// TIA Portal project "TestEssProtoFreia" (V13)

(* hardware
DEVICE "Station S7300/ET200M_1"  S7-300 station
   slot 0: "Châssis_0"  Rail  6ES7 390-1***0-0AA0
   slot 1: "Châssis_1"  Rail  6ES7 390-1***0-0AA0
   slot 1: "PS 307 2A_1"  PS 307 2A  6ES7 307-1BA01-0AA0
   slot 1: "PS 307 2A_1"  PS 307 2A  6ES7 307-1BA01-0AA0
   slot 2: "PLC_1"  CPU 315-2 DP  6ES7 315-2AH14-0AB0  V3.3
      slot 0: "Interface MPI_1"  MPI
      slot 1: "Interface DP_1"  DP
   slot 3: "IM 360_1"  6ES7 360-3AA01-0AA0
      slot 1: "Interface d'émission IM_1"  6ES7 360-3AA00-0AA0
   slot 3: "IM 361_1"  6ES7 361-3CA01-0AA0
      slot 1: "Interface d'émission IM_1"  6ES7 360-3AA00-0AA0
      slot 2: "Interface de réception IM_1"  6ES7 361-3CA00-0AA0
   slot 4: "DO 16x24VDC/0.5A_2"  DO16 x 24VDC / 0.5A  6ES7 322-1BH01-0AA0
   slot 4: "CP 343-1 Lean_1"  CP 343-1 LEAN  6GK7 343-1CX10-0XE0  V2.2
   slot 5: "DO 16x24VDC/0.5A_1"  DO16 x 24VDC / 0.5A  6ES7 322-1BH01-0AA0
   slot 5: "DI 16x24VDC_1"  DI16 x 24VDC  6ES7 321-1BH02-0AA0
   slot 6: "AI 8x12BIT_1"  AI8 x 12 bits  6ES7 331-7KF02-0AB0
   slot 6: "AI 8x12BIT_1"  AI8 x 12 bits  6ES7 331-7KF02-0AB0
   slot 7: "AI 8x12BIT_2"  AI8 x 12 bits  6ES7 331-7KF02-0AB0
   slot 7: "AO 8x12BIT_1"  AO8 x 12 bits  6ES7 332-5HF00-0AB0
   slot 8: "AI 8x12BIT_3"  AI8 x 12 bits  6ES7 331-7KF02-0AB0
   slot 8: "AO 4x12BIT_1"  AO4 x 12 bits  6ES7 332-5HD01-0AB0
   slot 9: "AI 8x16BIT_1"  AI8 x 16 bits  6ES7 331-7NF00-0AB0
   slot 9: "AO 4x12BIT_2"  AO4 x 12 bits  6ES7 332-5HD01-0AB0
DEVICE "Appareil GSD_1"  GSD.Device
   slot 0: "Châssis_0"  Rail
DEVICE "Appareil GSD_3"  GSD.Device
   slot 0: "Châssis_0"  Rail
DEVICE "Appareil GSD_4"  GSD.Device
   slot 0: "Châssis_0"  Rail
*)

// ===== PLC "PLC_1"  CPU 315-2 DP =====

VAR_GLOBAL   // PLC tag table "Table de variables standard"
   "TT_04" AT %ID720 : Real;
   "TT_218" AT %ID724 : Real;
   "TT_08CM" AT %ID728 : Real;
   "TT_217" AT %ID732 : Real;
   "TT_210" AT %ID736 : Real;
   "TT_209" AT %ID740 : Real;
   "TT_214" AT %ID744 : Real;
   "TT_03" AT %ID780 : Real;
   "TT_205" AT %ID784 : Real;
   "TT_05" AT %ID788 : Real;
   "TT_213" AT %ID792 : Real;
   "TT_14" AT %ID796 : Real;
   "TT_203" AT %ID800 : Real;
   "TT_204" AT %ID804 : Real;
   "TT_211" AT %ID808 : Real;
   "TT_202" AT %ID336 : Real;
   "TT_201" AT %ID340 : Real;
   "TT_104" AT %ID344 : Real;
   "TT_01CM" AT %ID348 : Real;
   "TT_115" AT %ID352 : Real;
   "TT_115bis" AT %ID356 : Real;
   "TT_208" AT %ID360 : Real;
   "TT_07" AT %ID364 : Real;
   "TT_12" AT %ID404 : Real;
   "TT_101" AT %ID408 : Real;
   "TT_103" AT %ID412 : Real;
   "TT_102" AT %ID416 : Real;
   "TT_04bis" AT %ID420 : Real;
   "TT_206" AT %ID424 : Real;
   "TT_02" AT %ID844 : Real;
   "TT_117" AT %ID856 : Real;
   "TT_106" AT %ID860 : Real;
   "TT_116" AT %ID864 : Real;
   "TT_118" AT %ID868 : Real;
   "TT_110" AT %ID872 : Real;
   "TT_207" AT %ID908 : Real;
   "TT_111" AT %ID924 : Real;
   "TT_107" AT %ID928 : Real;
   "TT_06" AT %ID932 : Real;
   "Tag_1" AT %IW3 : Word;
   "TimerDefauCom1" AT %T20 : Timer;
   "TimerDefauCom2" AT %T21 : Timer;
   "TT_215" AT %ID716 : Real;
   "CABTF4_voie10" AT %ID912 : Real;
   "CABTF4_voie11" AT %ID916 : Real;
   "CABTF4_voie12" AT %ID920 : Real;
   "Tag_45" AT %MD224 : Real;
   "Tag_46" AT %MW230 : Word;
   "Tag_47" AT %MW240 : Word;
   "Tag_48" AT %MD240 : Real;
   "Tag_49" AT %MD238 : DWord;
   "Tag_50" AT %MW238 : Word;
   "Tag_51" AT %MW242 : Word;
   "Tag_52" AT %MD244 : Real;
   "Tag_53" AT %IW388 : Int;
   "Tag_27" AT %MW600 : Word;
   "Tag_28" AT %MD602 : Real;
   "Tag_30" AT %M700.0 : Bool;
   "Tag_31" AT %M700.1 : Bool;
   "Tag_32" AT %M800.0 : Bool;
   "Tag_34" AT %MW804 : Int;
   "Tag_36" AT %MD808 : Real;
   "Tag_37" AT %MD812 : Real;
   "Tag_38" AT %MW816 : Word;
   "Tag_40" AT %M800.1 : Bool;
   "Tag_41" AT %M800.2 : Bool;
   "Tag_42" AT %MW802 : Int;
   "Tag_43" AT %MD804 : Real;
   "Tag_54" AT %MW820 : Word;
   "TT103_OHM" AT %MD820 : Real;
   "Tag_56" AT %IW646 : Word;
   "Tag_57" AT %IW648 : Word;
   "Tag_58" AT %IW480 : Word;
   "Tag_59" AT %IW482 : Word;
   "Tag_60" AT %IW472 : Word;
   "Tag_61" AT %IW474 : Word;
   "Tag_62" AT %IW464 : Word;
   "Tag_63" AT %IW466 : Word;
   "LocalMode" AT %M251.0 : Bool;
   "Tag_3" AT %M3.6 : Bool;
END_VAR

VAR_GLOBAL   // PLC tag table "Digital Input"
   "GV_70_CmInsulVacc:Open" AT %I0.0 : Bool;   // Cryomodule insulating vacuum Gate valve 70 open
   "GV_70_CmInsulVacc:Close" AT %I0.1 : Bool;   // Cryomodule insulating vacuum Gate valve 70 close
   "GV_71_CmInsulVacc:Open" AT %I0.3 : Bool;   // Cryomodule insulating vacuum Gate valve 71 open
   "GV_71_CmInsulVacc:Close" AT %I0.4 : Bool;   // Cryomodule insulating vacuum Gate valve 71 close
   "GV_72_VbInsulVacc:Open" AT %I0.6 : Bool;   // Cryomodule insulating vacuum Gate valve 72 open
   "GV_72_VbInsulVacc:Close" AT %I0.7 : Bool;   // Cryomodule insulating vacuum Gate valve 72 close
   "GV72_closed" AT %I1.1 : Bool;   // Cryomodule insulating vacuum Gate valve 72 closed
   "GV70_open" AT %I1.2 : Bool;   // Cryomodule insulating vacuum Gate valve 70 open
   "Tag_4" AT %I2.0 : Bool;
   "GV72_open" AT %I1.0 : Bool;   // Cryomodule insulating vacuum Gate valve 72 open
   "GV70_closed" AT %I1.3 : Bool;   // Cryomodule insulating vacuum Gate valve 70 closed
   "RV90_open" AT %I1.4 : Bool;   // He release valve
   "RV90_closed" AT %I1.5 : Bool;   // He release valve
END_VAR

VAR_GLOBAL   // PLC tag table "analog output"
   "CMD_CV_01" AT %QW384 : Int;
   "CMD_CV_02" AT %QW386 : Int;
   "CMD_CV_03" AT %QW388 : Int;
   "CMD_CV_04" AT %QW390 : Int;
   "CMD_CV_05" AT %QW392 : Int;
   "CMD_CV_07" AT %QW394 : Int;
   "CMD_CV_60" AT %QW396 : Int;
   "CMD_CV_61" AT %QW398 : Int;
   "CMD_CV_62" AT %QW400 : Int;
   "Sana_ASCO_1" AT %QW402 : Int;
   "Sana_ASCO_2" AT %QW404 : Int;
END_VAR

VAR_GLOBAL   // PLC tag table "mem"
   "always_1" AT %M0.1 : Bool;
   "always_0" AT %M0.0 : Bool;
   "unscal_ret_val" AT %MW40 : Word;
   "CV01_HMI_VAL" AT %MD4 : Real;
   "CV02_HMI_VAL" AT %MD8 : Real;
   "CV03_HMI_VAL" AT %MD12 : Real;
   "CV04_HMI_VAL" AT %MD16 : Real;
   "CV05_HMI_VAL" AT %MD20 : Real;
   "CV07_HMI_VAL" AT %MD24 : Real;
   "CV60_HMI_VAL" AT %MD28 : Real;
   "CV61_HMI_VAL" AT %MD36 : Real;
   "unscal_ret_val_1" AT %MW42 : Word;
   "unscal_ret_val_2" AT %MW44 : Word;
   "unscal_ret_val_3" AT %MW46 : Word;
   "unscal_ret_val_4" AT %MW48 : Word;
   "unscal_ret_val_5" AT %MW50 : Word;
   "unscal_ret_val_6" AT %MW52 : Word;
   "unscal_ret_val_7" AT %MW54 : Word;
   "unscal_ret_val_8" AT %MW56 : Word;
   "CV62_HMI_VAL" AT %MD32 : Real;
   "Tag_7" AT %MD701 : Real;
   "Tag_8" AT %MD706 : Real;
   "Tag_9" AT %MD710 : Real;
   "Tag_10" AT %MD714 : Real;
   "Tag_11" AT %MD718 : Real;
   "Tag_12" AT %MD722 : Real;
   "Tag_13" AT %MD726 : Real;
   "Tag_14" AT %MD730 : Real;
   "Tag_15" AT %MD734 : Real;
   "Tag_16" AT %MW100 : Word;
   "Tag_17" AT %MW102 : Word;
   "Tag_18" AT %MW104 : Word;
   "Tag_19" AT %MW106 : Word;
   "Tag_20" AT %MW108 : Word;
   "Tag_21" AT %MW110 : Word;
   "Tag_22" AT %MW112 : Word;
   "Tag_23" AT %MW114 : Word;
   "Tag_24" AT %MW116 : Word;
   "TT670_(OHMS)" AT %MD58 : Real;
   "LT03_DepHaut" AT %M0.3 : Bool;
   "LT03_DepBas" AT %M0.4 : Bool;
   "LT03_DefSond" AT %M0.5 : Bool;
   "LT03_TypeDef" AT %MW66 : Int;
   "LT03_ValMax" AT %MD72 : Real;
   "LT03_ValMin" AT %MD76 : Real;
   "LT03_NiveauHel" AT %MD80 : Real;
   "CV02_ManAuto" AT %M0.6 : Bool;
   "CV03_ManAuto" AT %M0.7 : Bool;
   "CV61_ManAuto" AT %M1.0 : Bool;
   "ScaleErreurPT60" AT %MW68 : Word;
   "ScaleErreurPT01" AT %MW88 : Word;
   "ScaleErreurVidePT73" AT %MW90 : Word;
   "VidePT73Tension" AT %MD92 : Real;
   "CV01PosInit" AT %M1.1 : Bool;
   "CV02PosInit" AT %M1.2 : Bool;
   "CV03PosInit" AT %M1.3 : Bool;
   "CV04PosInit" AT %M1.4 : Bool;
   "CV05PosInit" AT %M1.5 : Bool;
   "CV07PosInit" AT %M1.6 : Bool;
   "CV60PosInit" AT %M1.7 : Bool;
   "CV61PosInit" AT %M62.0 : Bool;
   "CV62PosInit" AT %M62.1 : Bool;
   "CmdVanneEtatInitial" AT %M62.2 : Bool;
   "VanneEnPositionInitial" AT %M62.3 : Bool;
   "CmdVanneEtatCdt" AT %M62.4 : Bool;
   "Etat initial" AT %M62.5 : Bool;
   "CV01PosCdt" AT %M62.6 : Bool;
   "CV02PosCdt" AT %M62.7 : Bool;
   "CV03PosCdt" AT %M63.0 : Bool;
   "CV04PosCdt" AT %M63.1 : Bool;
   "CV05PosCdt" AT %M63.2 : Bool;
   "CV07PosCdt" AT %M63.3 : Bool;
   "CV60PosCdt" AT %M63.4 : Bool;
   "CV61PosCdt" AT %M63.5 : Bool;
   "CV62PosCdt" AT %M63.6 : Bool;
   "VanneEnPositionCdt" AT %M63.7 : Bool;
   "EtatCdtCryo" AT %M64.0 : Bool;
   "ScaleErreurVidePT71" AT %MW96 : Word;
   "VidePT71Tension" AT %MD118 : Real;
   "AutorizationMefAzote" AT %M64.1 : Bool;
   "ReguleCV61ON" AT %M64.2 : Bool;
   "CmdVanneEtatMEFazote" AT %M64.3 : Bool;
   "CmdVanneEtatMEFhelium" AT %M64.4 : Bool;
   "EtatMEFhelium" AT %M64.5 : Bool;
   "LT01_NiveauHel" AT %MD122 : Real;
   "LT01_DepHaut" AT %M64.6 : Bool;
   "LT01_DepBas" AT %M64.7 : Bool;
   "LT01_DefSond" AT %M65.0 : Bool;
   "LT01_TypeDef" AT %MW98 : Int;
   "LT01_ValMax" AT %MD126 : Real;
   "LT01_ValMin" AT %MD130 : Real;
   "EtatModeStandBy" AT %M65.1 : Bool;
   "NumEtape" AT %MW134 : Int;
   "EtatMode2K" AT %M65.2 : Bool;
   "EtatAttMef" AT %M65.3 : Bool;
   "EtatMEFazote" AT %M65.4 : Bool;
   "CdtInfraErreur" AT %M65.5 : Bool;
   "CdtInfraOk" AT %M65.6 : Bool;
   "DmdMefAzote" AT %M65.7 : Bool;
   "DmdMefHelium" AT %M136.0 : Bool;
   "DmdMode2K" AT %M136.1 : Bool;
   "DmdArretMode2k" AT %M136.2 : Bool;
   "DmdModeStandby" AT %M136.3 : Bool;
   "DmdArretModeStandby" AT %M136.4 : Bool;
   "TransMode4K" AT %M136.5 : Bool;
   "EtatMode4k" AT %M136.6 : Bool;
   "DesactiveGraph" AT %M136.7 : Bool;
   "MettreEtatInitial" AT %M137.0 : Bool;
   "AcquitterErreurGraph" AT %M137.1 : Bool;
   "Graph/manuelle" AT %M137.2 : Bool;
   "ErreurSupervision" AT %M137.3 : Bool;
   "conditionTempMEFheliumOK" AT %M137.4 : Bool;
   "tt77h" AT %M137.6 : Bool;
   "tt77l" AT %M137.7 : Bool;
   "tt77alm" AT %M140.0 : Bool;
   "tt77typedef" AT %MW142 : Int;
   "tt77max" AT %MD144 : Real;
   "tt77min" AT %MD148 : Real;
   "OB32_year" AT %MB152 : Byte;
   "SeuilHautPressionBoteil" AT %MD156 : Real;
   "DmdChangementBouteil" AT %M140.1 : Bool;
   "Tag_M" AT %M140.2 : Bool;
   "FCtoDBok" AT %M140.3 : Bool;
   "unscal_ret_val_asco_1" AT %MW160 : Word;
   "unscal_ret_val_asco_2" AT %MW162 : Word;
   "ASCO1PosInit" AT %M140.4 : Bool;
   "ASCO2PosInit" AT %M140.5 : Bool;
   "ASCO1PosCdt" AT %M140.6 : Bool;
   "ASCO2PosCdt" AT %M140.7 : Bool;
   "RéguleASCO02_SP" AT %MD168 : Real;
   "ASCOenManuel" AT %M141.0 : Bool;
   "Asco02ManValeur" AT %MD176 : Real;
   "PositionASCO02" AT %MD186 : Real;
   "CV01_2K_MAN_value" AT %MD192 : Real;
   "NiveauHel_Hmi" AT %MD196 : Real;
   "Etatrechauffage" AT %M141.2 : Bool;
   "TriggerPIDcv03" AT %MD200 : Real;
   "LT03LevelSP" AT %MD204 : Real;
   "TriggerPIDcv02" AT %MD208 : Real;
   "LT01LevelSP" AT %MD212 : Real;
   "TriggerPIDcv01" AT %MD216 : Real;
   "LT01LevelSP2k" AT %MD220 : Real;
   "CmdVanneEtatstdby" AT %M141.3 : Bool;
   "CV60_ManAuto" AT %M141.4 : Bool;
   "CV07_ManAuto" AT %M141.5 : Bool;
   "CV04_ManAuto" AT %M141.6 : Bool;
   "CV01_ManAuto" AT %M141.7 : Bool;
   "ScaleErreurPressionDiff" AT %MW224 : Word;
   "Tag_26" AT %MW190 : Word;
   "Tag_6" AT %MD746 : Real;
   "Scale_erreur_tt670" AT %MW2 : Word;
   "TT_001:OHMS" AT %MD84 : Real;
   "INIT" AT %M0.2 : Bool;
   "ScaleErreurNiveauBouteil" AT %MW226 : Word;
   "LT01RegActive" AT %M230.0 : Bool;
   "LT03RegActive" AT %M230.1 : Bool;
   "LT01Reg2KActive" AT %M230.2 : Bool;
   "StartHeating" AT %M138.0 : Bool;
   "StopHeating" AT %M138.1 : Bool;
   "point1sec" AT %M300.0 : Bool;
   "point1secPls" AT %M301.0 : Bool;
   "point1secMem" AT %M302.0 : Bool;
   "oneSec" AT %M300.5 : Bool;
   "oneSecPls" AT %M301.5 : Bool;
   "oneSecMem" AT %M302.5 : Bool;
   "HNOSS_COMM_OK" AT %M138.2 : Bool;
   "Separators_empty" AT %M137.5 : Bool;
   "Ret_val" AT %MW164 : Int;
   "OB32_month" AT %MB153 : Byte;
   "OB32_day" AT %MB154 : Byte;
   "OB32_hour" AT %MB155 : Byte;
   "OB32_min" AT %MB156 : Byte;
   "OB32_sec" AT %MB157 : Byte;
   "OB32_ms_dow" AT %MW158 : Word;
   "OneMinute" AT %M231.0 : Bool;
   "Tag_2" AT %MD306 : Real;
   "Minute_mem" AT %MB160 : Byte;   // A help variable to store the previous readout
   "OneMinute_CV03_mem" AT %M3.0 : Bool;   // Memory bit for positive pulse used in the control of
   "OnOff_test" AT %M3.1 : Bool;   // A bit for temporary tests (debugging)
   "2KModeStart_mem" AT %M3.2 : Bool;
   "OneMinute_CV01_mem" AT %M3.3 : Bool;
   "WarmUpStart_mem" AT %M3.4 : Bool;
   "LT02_NiveauHel" AT %MD180 : Real;
   "LT02_TypeDef" AT %MW166 : Int;
   "LT02_DefSond" AT %M70.0 : Bool;
   "LT02_DepBas" AT %M70.1 : Bool;
   "LT02_DepHaut" AT %M70.2 : Bool;
   "LT02_ValMin" AT %MD172 : Real;
   "LT02_ValMax" AT %MD232 : Real;
   "INH_BIT" AT %M3.5 : Bool;
END_VAR

VAR_GLOBAL CONSTANT   // PLC tag table "mem"
   "m16.0" : Bool := 1;
END_VAR

VAR_GLOBAL   // PLC tag table "analog input"
   "RetourPositionCV01" AT %IW288 : Int;
   "RetourPositionCV02" AT %IW290 : Int;
   "RetourPositionCV03" AT %IW292 : Int;
   "RetourPositionCV04" AT %IW294 : Int;
   "RetourPositionCV05" AT %IW296 : Int;
   "RetourPositionCV07" AT %IW298 : Int;
   "RetourPositionCV60" AT %IW300 : Int;
   "RetourPositionCV61" AT %IW302 : Int;
   "RetourPositionCV62" AT %IW304 : Int;
   "Eana_NiveauH_LT03" AT %IW306 : Int;
   "Eana_VidePT75" AT %IW320 : Int;   // TEMPERATURE PT100
   "Eana_PressionPT60" AT %IW312 : Int;
   "Eana_PressionPT01" AT %IW314 : Int;
   "Eana_VidePT71" AT %IW316 : Int;
   "Eana_VidePT73" AT %IW318 : Int;
   "Eana_NiveauH_LT01" AT %IW308 : Int;
   "Eana_NiveauH_LT02" AT %IW310 : Int;
   "Eana_VidePT77" AT %IW322 : Int;
   "TT_109" AT %ID400 : Real;
   "TT_105" AT %ID428 : Real;
   "TT_02JM" AT %ID586 : DWord;
   "TT_03JM" AT %ID590 : DWord;
   "TT_04JM" AT %ID594 : DWord;
   "TT_09" AT %ID598 : DWord;
   "TT_10" AT %ID602 : DWord;
   "Eana_TT77_ohm" AT %IW328 : Int;   // 4 fils
   "Eana_ASCO2" AT %IW324 : Int;
   "Eana_PressionDiff" AT %IW326 : Int;
   "TT_01" AT %ID518 : DWord;
   "TT_08" AT %ID522 : DWord;
   "TT_91" AT %ID526 : DWord;
   "TT_92" AT %ID530 : DWord;
   "TT_93" AT %ID534 : DWord;
   "TT_94" AT %ID538 : DWord;
   "TT_95" AT %ID542 : DWord;
   "TT_97" AT %ID546 : DWord;
   "TT_98" AT %ID582 : DWord;
   "TT120" AT %IW488 : Int;
   "FT11" AT %IW332 : Int;   // Mass Flowmeter 0-150 mg/s Coupler 1
   "FT21" AT %IW334 : Int;   // Mass Flowmeter 0-150 mg/s Coupler 2
   "TT110" AT %IW496 : Int;   // Thermocouple with 4-20mA adapter
   "TT210" AT %IW498 : Int;   // Thermocouple with 4-20mA adapter
   "TT220" AT %IW492 : Int;
   "PT02_direct" AT %IW654 : Int;
END_VAR

VAR_GLOBAL   // PLC tag table "Digital output"
   "voie 1 chaufferette BV" AT %Q72.0 : Bool;
   "voie 2 chaufferette BV" AT %Q72.1 : Bool;
   "voie 3 chaufferette BV" AT %Q72.2 : Bool;
   "voie 4 chaufferette BV" AT %Q72.3 : Bool;
   "voie 5 chaufferette BV" AT %Q72.4 : Bool;
   "voie 6 chaufferette BV" AT %Q72.5 : Bool;
   "voie 7 chaufferette BV" AT %Q72.6 : Bool;
   "voie 8 chaufferette BV" AT %Q72.7 : Bool;
   "voie 9 chaufferette BV" AT %Q73.0 : Bool;
   "voie 1 chaufferette CM" AT %Q20.2 : Bool;
   "voie 2 chaufferette CM" AT %Q20.3 : Bool;
   "voie 3 chaufferette CM" AT %Q20.4 : Bool;
   "voie 4 chaufferette CM" AT %Q20.5 : Bool;
   "voie 5 chaufferette CM" AT %Q20.6 : Bool;
   "voie 6 chaufferette CM" AT %Q20.7 : Bool;
   "voie 8 chaufferette CM" AT %Q21.1 : Bool;
   "voie 10  chaufferette BV" AT %Q73.1 : Bool;
   "voie 11 chaufferette BV" AT %Q73.2 : Bool;
   "voie 7 chaufferette CM" AT %Q21.0 : Bool;
   "GV72_OpenCmd" AT %Q20.0 : Bool;
   "RV90_OpenCmd" AT %Q20.1 : Bool;
   "voie 9 chaufferette CM" AT %Q21.2 : Bool;
   "voie 10 chaufferette CM" AT %Q21.3 : Bool;
   "voie 11 chaufferette CM" AT %Q21.4 : Bool;
   "voie 12 chaufferette CM" AT %Q21.5 : Bool;
   "EH12 Cpl1" AT %Q21.6 : Bool;
   "EH22 Cpl2" AT %Q21.7 : Bool;
   "CM_CryoOK" AT %Q73.7 : Bool;   // Interlock signal for RF slow interlock
   "GV70_OpenCmd" AT %Q73.6 : Bool;
END_VAR

VAR_GLOBAL   // PLC tag table "EPICS_comm"
   "RCV_NDR" AT %M250.3 : Bool;
   "RCV_ERR" AT %M250.4 : Bool;
   "RECV_status" AT %MW254 : Word;
   "RECV_len" AT %MW256 : Int;
   "EPICS_send_T1" AT %T1 : Timer;
   "EPICS_do_send" AT %M250.0 : Bool;
   "EPICS_send_T0" AT %T0 : Timer;
   "SND_DONE" AT %M250.1 : Bool;
   "SND_ERR" AT %M250.2 : Bool;
   "SEND_status" AT %MW252 : Word;
   "ACT_SEND" AT %M250.5 : Bool;
   "SND_BUSY" AT %M250.6 : Bool;
   "SND_CLK_RLO_MEM" AT %M250.7 : Bool;
   "SND_STAT_SAVE" AT %MW258 : Word;
   "RCV_STAT_SAVE" AT %MW260 : Word;
   "RCV_CNT" AT %C1 : Counter;
   "EPICS_COMM_OK" AT %M270.0 : Bool;
   "SND_DONE(1)" AT %M270.1 : Bool;
   "SND_ERR(1)" AT %M270.2 : Bool;
   "RCV_NDR(1)" AT %M270.3 : Bool;
   "RCV_ERR(1)" AT %M270.4 : Bool;
   "ACT_SEND(1)" AT %M270.5 : Bool;
   "SND_BUSY(1)" AT %M270.6 : Bool;
   "SND_CLK_RLO_MEM(1)" AT %M270.7 : Bool;
   "SEND_status(1)" AT %MW272 : Word;
   "RECV_status(1)" AT %MW274 : Word;
   "RECV_len(1)" AT %MW276 : Int;
   "SND_STAT_SAVE(1)" AT %MW278 : Word;
   "RCV_STAT_SAVE(1)" AT %MW280 : Word;
END_VAR

TYPE "FValve_cmd"
   STRUCT
      cmdOpen : Bool;
      cmdClose : Bool;
      cmdAuto : Bool;
      cmdMan : Bool;
   END_STRUCT;
END_TYPE

TYPE "Cernox"
   STRUCT
      board1 : Array[0..7] of Real;
      board2 : Array[0..7] of Real;
      stat : Array[0..3] of Word;
   END_STRUCT;
END_TYPE

TYPE "FValve_s"
   STRUCT
      sOpen : Bool;
      sClosed : Bool;
      sCmdOpen : Bool;
      sAuto : Bool;
      sFault : Bool;
   END_STRUCT;
END_TYPE

TYPE "CV_stat"
   STRUCT
      sRdV : Real;
      sSetV : Real;
      sSetVAuto : Real;
      sAuto : Bool;
      sPosInit : Bool;
      sPosCnd : Bool;
   END_STRUCT;
END_TYPE

TYPE "CV_cmd"
   STRUCT
      cSetv : Real;
      cmdMan : Bool;
      cmdAuto : Bool;
      cmdSet : Bool;
   END_STRUCT;
END_TYPE

TYPE "EH_cmd"
   STRUCT
      cmdAuto : Bool;
      cmdMan : Bool;
      cmdSet : Bool;
      cmdRst : Bool;
      cmdHL : Bool;
      cmdLL : Bool;
      cHL : Real;
      cLL : Real;
   END_STRUCT;
END_TYPE

TYPE "EH_stat"
   STRUCT
      sAuto : Bool;
      sTsw : Bool;
      sCmd : Bool;
      sCmdAuto : Bool;
      sHtrOn : Bool;
      sHL : Real;
      sLL : Real;
   END_STRUCT;
END_TYPE

TYPE "Real_val_cmd"
   STRUCT
      cmdSet : Bool;
      cSetV : Real;
   END_STRUCT;
END_TYPE

TYPE "Real_val_stat"
   STRUCT
      sSetV : Real;
   END_STRUCT;
END_TYPE

TYPE "LevelMeter"
   STRUCT
      Level : Real;
      Visu : Int;
      SensorFlt : Bool;
      OverRange : Bool;
      UnderRange : Bool;
   END_STRUCT;
END_TYPE

TYPE "UDT_HEATER"
VERSION : 0.1
   STRUCT
      XH : Bool;
      X : Bool;
      H : Bool;
      Raz_Fct_Run : Bool;
      Ok : Bool;
      Pilot : Bool;
      R_EH : Bool;
      TS_Calc : Bool;
      TS : Bool;
      Pilot_Calc : Bool;
      R_ExtCmd : Bool;
      Not_Connected : Bool;
      P_TS_Ton : DInt;
      TS_Ton : DInt;
      P_TS_Toff : DInt;
      TS_Toff : DInt;
      T_run : DInt;
      Tt_Max : Real;
      Tt_Min : Real;
      ValueA : Real;
      ValueB : Real;
      ValueC : Real;
      ValueD : Real;
      ValueE : Real;
      ValueF : Real;
      Nb_Tt : Int;
      P_Pilot_Ton : DInt;
      Pilot_Ton : DInt;
   END_STRUCT;
END_TYPE

TYPE "Epi_to_Plc_Valve"
VERSION : 0.0
   STRUCT
      cmdAuto : Bool;
      cmdMan : Bool;
      cmdSet : Bool;
      cmdRst : Bool;
      cmdAck : Bool;
      cmdSimSet : Bool;
      cmdSimRst : Bool;
   END_STRUCT;
END_TYPE

TYPE "Plc_to_Epi_Valve"
VERSION : 0.0
   STRUCT
      sAuto : Bool;
      sSim : Bool;
      sCmd : Bool;
      sOn : Bool;
      sOff : Bool;
      sNO : Bool;
      sOnFlt : Bool;
      sOffFlt : Bool;
      sFlt : Bool;
      sCmdAuto : Bool;
   END_STRUCT;
END_TYPE

TYPE "UDT_VALVES"
VERSION : 0.1
   STRUCT
      XH : Bool;
      X : Bool;
      H : Bool;
      Ack : Bool;
      Inh : Bool;
      Raz_Fct_Run : Bool;
      Ok : Bool;
      Df : Bool;
      Df_on : Bool;
      Df_off : Bool;
      Rzson : Bool;
      Rzsoff : Bool;
      R_in : Bool;
      R_out : Bool;
      Rxv : Bool;
      Not_Connected : Bool;
      T_run : DInt;
      C_run : DInt;
      Gen : Struct
      END_STRUCT;
      Internal : Struct
      END_STRUCT;
   END_STRUCT;
END_TYPE

DATA_BLOCK "Pression"   // DB10
{ S7_Optimized_Access := 'FALSE' }
VERSION : 0.1
   VAR
      PressionPT60_Val : Real;
      PressionPT01_Val : Real;
      PressionVidePT73 : Real;
      PressionVidePT71 : Real;
      PT02_direct : Real;
      NiveauHeBV : Real;
      NiveauHeCM : Real;
      PressionDiff : Real;
      NiveauBouteilHe : Real;
      PressionVidePT75 : Real;
      PressionVidePT77 : Real;
      temp_bride_coupleur : Real;
   END_VAR
BEGIN
END_DATA_BLOCK

DATA_BLOCK "ReceivePT100"   // DB11
{ S7_Optimized_Access := 'FALSE' }
VERSION : 0.1
   VAR
      "TT77_(K)" : Real;
      "TT77_(R)" : Real;
      "TT03_(K)" : Real;
      "TTxx_(K)" : Real;
      "TTyy_(K)" : Real;
   END_VAR
BEGIN
END_DATA_BLOCK

DATA_BLOCK "graf_DB"   // DB13
{ S7_Optimized_Access := 'FALSE' }
VERSION : 0.1
// stored: InstanceOfName graf
"graf"
BEGIN
END_DATA_BLOCK

DATA_BLOCK "Position_vannes"   // DB15
{ S7_Optimized_Access := 'FALSE' }
VERSION : 0.1
   VAR
      PositionCV01 : Real;
      PositionCV02 : Real;
      PositionCV03 : Real;
      PositionCV04 : Real;
      PositionCV05 : Real;
      PositionCV07 : Real;
      PositionCV60 : Real;
      PositionCV61 : Real;
   END_VAR
BEGIN
END_DATA_BLOCK

DATA_BLOCK "PLC_to_Epics"   // DB100
{ S7_Optimized_Access := 'FALSE' }
VERSION : 0.1
   VAR
      sLocal : Bool;
      sManual : Bool;
      sGrafcetERR : Bool;
      sGS1 : Bool;
      sGS2 : Bool;
      sGS3 : Bool;
      sGS4 : Bool;
      sGS5 : Bool;
      sGS6 : Bool;
      sGS7 : Bool;
      sGS8 : Bool;
      sGS10 : Bool;
      sTransTempOK : Bool;
      sTransMode4K : Bool;
      CV550_PID_on : Bool;
      CV60_PID_on : Bool;
      CV01_PID_on : Bool;
      CV02_PID_on : Bool;
      CV03_PID_on : Bool;
      EpicsCommOK : Bool;
      HNOSSCommOK : Bool;
      CV5202_OpenReq : Bool;
      General : Array[0..15] of Real;
      CABTF1 : "Cernox";
      CABTF2 : "Cernox";
      CABTF3 : "Cernox";
      CABTF_spare : "Cernox";
      CV01 : "CV_stat";
      CV02 : "CV_stat";
      CV03 : "CV_stat";
      CV04 : "CV_stat";
      CV05 : "CV_stat";
      CV07 : "CV_stat";
      CV60 : "CV_stat";
      CV61 : "CV_stat";
      CV62 : "CV_stat";
      CV550 : "CV_stat";
      CV551 : "CV_stat";
      CV552 : "CV_stat";
      CVRes01 : "CV_stat";
      CVRes02 : "CV_stat";
      EH90 : "EH_stat";
      "EH93-96" : "EH_stat";
      "EH63-70" : "EH_stat";
      "EH61-62" : "EH_stat";
      "EH60_67-69" : "EH_stat";
      "EH97-98" : "EH_stat";
      "spare-VB-7" : "EH_stat";
      "spare-VB-8" : "EH_stat";
      "spare-VB-9" : "EH_stat";
      "spare-VB-10" : "EH_stat";
      "spare-VB-11" : "EH_stat";
      EH01 : "EH_stat";
      EH02 : "EH_stat";
      EH10 : "EH_stat";
      EH20 : "EH_stat";
      "spare-CM-5" : "EH_stat";
      "spare-CM-6" : "EH_stat";
      "spare-CM-7" : "EH_stat";
      "spare-CM-8" : "EH_stat";
      "spare-CM-9" : "EH_stat";
      "spare-CM-10" : "EH_stat";
      "spare-CM-11" : "EH_stat";
      "spare-CM-12" : "EH_stat";
      EH12 : "EH_stat";
      EH22 : "EH_stat";
      "EH-Res" : Array[0..6] of "EH_stat";
      FV101 : "FValve_s";
      FV102 : "FValve_s";
      LT01 : "LevelMeter";
      LT03 : "LevelMeter";
      PT60 : Real;
      PT01 : Real;
      PT73 : Real;
      PT71 : Real;
      PT75 : Real;
      PT77 : Real;
      TrigPID_CV01 : "Real_val_stat";
      PID_LT01_CV01_SP : "Real_val_stat";
      TrigPID_CV02 : "Real_val_stat";
      PID_LT01_CV02_SP : "Real_val_stat";
      TrigPID_CV03 : "Real_val_stat";
      PID_LT03_CV03_SP : "Real_val_stat";
      PID_PT01_CV550_SP : "Real_val_stat";
      TT77 : "LevelMeter";
      PT04 : Real;
      FT11 : "LevelMeter";
      FT21 : "LevelMeter";
      TT110 : "LevelMeter";
      TT210 : "LevelMeter";
      TT120 : "LevelMeter";
      TT220 : "LevelMeter";
      S5_P_FT552_MIN_GB : "Real_val_stat";
      S5_P_FT552_MAX_GB : "Real_val_stat";
      S5_P_FT552_MIN_C : "Real_val_stat";
      S5_P_FT552_MAX_C : "Real_val_stat";
      S4step : Byte;
      S5step : Byte;
      S6step : Byte;
      S7step : Byte;
      S8step : Byte;
      S9step : Byte;
      S10step : Byte;
      SXstep : Byte;
      S8_P_CV01 : "Real_val_stat";
      LT02 : "LevelMeter";
      GV72 : "Plc_to_Epi_Valve";
      RV90 : "Plc_to_Epi_Valve";
      GV70 : "Plc_to_Epi_Valve";
      GV_spare1 : "Plc_to_Epi_Valve";
      CV01_PID_GAIN : "Real_val_stat";
      CV01_PID_TI : "Real_val_stat";
      CV01_PID_TD : "Real_val_stat";
      CV01_PID_TM_LAG : "Real_val_stat";
      CV02_PID_GAIN : "Real_val_stat";
      CV02_PID_TI : "Real_val_stat";
      CV02_PID_TD : "Real_val_stat";
      CV02_PID_TM_LAG : "Real_val_stat";
      CV03_PID_GAIN : "Real_val_stat";
      CV03_PID_TI : "Real_val_stat";
      CV03_PID_TD : "Real_val_stat";
      CV03_PID_TM_LAG : "Real_val_stat";
      CV60_PID_GAIN : "Real_val_stat";
      CV60_PID_TI : "Real_val_stat";
      CV60_PID_TD : "Real_val_stat";
      CV60_PID_TM_LAG : "Real_val_stat";
      PID_TT77_CV60_SP : "Real_val_stat";
      PT02_direct : Real;
      S8_P_CV01_Step7 : "Real_val_stat";
      dummy : Array[0..437] of Word;
   END_VAR
BEGIN
END_DATA_BLOCK

DATA_BLOCK "Epics_to_PLC"   // DB101
{ S7_Optimized_Access := 'FALSE' }
VERSION : 0.1
   VAR
      cmdLocalMode : Bool;
      cmdRemoteMode : Bool;
      cmdAutoMode : Bool;
      cmdManMode : Bool;
      cmdGrafcetInit : Bool;
      cmdGrafcetErrRst : Bool;
      cmdStartConditioning : Bool;
      cmdCondOK : Bool;
      cmdCondERR : Bool;
      cmdStartLN2cooling : Bool;
      cmdStartLHecooling : Bool;
      cmdStart2Kmode : Bool;
      cmdStop2Kmode : Bool;
      cmdStartSTBYmode : Bool;
      cmdStopSTBYmode : Bool;
      cmdStartHeating : Bool;
      cmdStopHeating : Bool;
      cmdAckn : Bool;
      TTxx : Real;
      TTyy : Real;
      General : Array[0..13] of DWord;
      CV01 : "CV_cmd";
      CV02 : "CV_cmd";
      CV03 : "CV_cmd";
      CV04 : "CV_cmd";
      CV05 : "CV_cmd";
      CV07 : "CV_cmd";
      CV60 : "CV_cmd";
      CV61 : "CV_cmd";
      CV62 : "CV_cmd";
      CV550 : "CV_cmd";
      CV551 : "CV_cmd";
      CV552 : "CV_cmd";
      CVRes01 : "CV_cmd";
      CVRes02 : "CV_cmd";
      EH90 : "EH_cmd";
      "EH93-96" : "EH_cmd";
      "EH63-70" : "EH_cmd";
      "EH61-62" : "EH_cmd";
      "EH60_67-69" : "EH_cmd";
      "EH97-98" : "EH_cmd";
      "spare-VB-7" : "EH_cmd";
      "spare-VB-8" : "EH_cmd";
      "spare-VB-9" : "EH_cmd";
      "spare-VB-10" : "EH_cmd";
      "spare-VB-11" : "EH_cmd";
      EH01 : "EH_cmd";
      EH02 : "EH_cmd";
      EH10 : "EH_cmd";
      EH20 : "EH_cmd";
      "spare-CM-5" : "EH_cmd";
      "spare-CM-6" : "EH_cmd";
      "spare-CM-7" : "EH_cmd";
      "spare-CM-8" : "EH_cmd";
      "spare-CM-9" : "EH_cmd";
      "spare-CM-10" : "EH_cmd";
      "spare-CM-11" : "EH_cmd";
      "spare-CM-12" : "EH_cmd";
      EH12 : "EH_cmd";
      EH22 : "EH_cmd";
      "EH-Res" : Array[0..6] of "EH_cmd";
      TrigPID_CV01 : "Real_val_cmd";
      PID_LT01_CV01_SP : "Real_val_cmd";
      TrigPID_CV02 : "Real_val_cmd";
      PID_LT01_CV02_SP : "Real_val_cmd";
      TrigPID_CV03 : "Real_val_cmd";
      PID_LT03_CV03_SP : "Real_val_cmd";
      PID_PT01_CV550_SP : "Real_val_cmd";
      S5_P_FT552_MIN_GB : "Real_val_cmd";
      S5_P_FT552_MAX_GB : "Real_val_cmd";
      S5_P_FT552_MIN_C : "Real_val_cmd";
      S5_P_FT552_MAX_C : "Real_val_cmd";
      S8_P_CV01 : "Real_val_cmd";
      GV72 : "Epi_to_Plc_Valve";
      RV90 : "Epi_to_Plc_Valve";
      GV70 : "Epi_to_Plc_Valve";
      GV_spare1 : "Epi_to_Plc_Valve";
      CV01_PID_GAIN : "Real_val_cmd";
      CV01_PID_TI : "Real_val_cmd";
      CV01_PID_TD : "Real_val_cmd";
      CV01_PID_TM_LAG : "Real_val_cmd";
      CV02_PID_GAIN : "Real_val_cmd";
      CV02_PID_TI : "Real_val_cmd";
      CV02_PID_TD : "Real_val_cmd";
      CV02_PID_TM_LAG : "Real_val_cmd";
      CV03_PID_GAIN : "Real_val_cmd";
      CV03_PID_TI : "Real_val_cmd";
      CV03_PID_TD : "Real_val_cmd";
      CV03_PID_TM_LAG : "Real_val_cmd";
      CV60_PID_GAIN : "Real_val_cmd";
      CV60_PID_TI : "Real_val_cmd";
      CV60_PID_TD : "Real_val_cmd";
      CV60_PID_TM_LAG : "Real_val_cmd";
      PID_TT77_CV60_SP : "Real_val_cmd";
      S8_P_CV01_Step7 : "Real_val_cmd";
      data : Array[0..84] of Real;
   END_VAR
BEGIN
END_DATA_BLOCK

DATA_BLOCK "Data_from_HNOSS"   // DB102
{ S7_Optimized_Access := 'FALSE' }
VERSION : 0.1
// Placeholder for data received from HNOSS
   VAR
      HeartBeat : Word;
      CV5202_PercOut : Real;
      CV5202_Open : Bool;
      CV5202_VALID : Bool;
      FV401_Closed : Bool;
      FV401_Open : Bool;
      FV501_Closed : Bool;
      FV501_Open : Bool;
      FV550_Closed : Bool;
      FV550_Open : Bool;
      FV551_Closed : Bool;
      FV551_Open : Bool;
      FV552_Closed : Bool;
      FV552_Open : Bool;
      FV553_Closed : Bool;
      FV553_Open : Bool;
      FV554_Closed : Bool;
      FV554_Open : Bool;
      FV555_Closed : Bool;
      FV555_Open : Bool;
      FT550 : Real;
      FT551 : Real;
      FT552 : Real;
      CV550 : Real;
      CV551 : Real;
      CV552 : Real;
      SQ9_state : Int;
      spare : Array[0..61] of Word;
   END_VAR
BEGIN
END_DATA_BLOCK

DATA_BLOCK "Data_to_HNOSS"   // DB103
{ S7_Optimized_Access := 'FALSE' }
VERSION : 0.1
// Data to be read by HNOSS
   VAR
      HeartBeat : Word;
      InitState : Bool;
      Conditioning : Bool;
      Purged : Bool;
      ScreenCooling : Bool;
      LHeCooling : Bool;
      Operation4K : Bool;
      Operation2K : Bool;
      Standby : Bool;
      WarmUp : Bool;
      RegOnMKS1 : Bool;
      RegOnMKS2 : Bool;
      RegOnMKS3 : Bool;
      SP_PT01_MKS2 : Real;
      CV550_MKS2 : Real;
      S4step : Byte;
      S5step : Byte;
      S6step : Byte;
      S7step : Byte;
      S8step : Byte;
      S9step : Byte;
      S10step : Byte;
      SXstep : Byte;
      spare : Array[0..139] of Byte;
   END_VAR
BEGIN
END_DATA_BLOCK

DATA_BLOCK "PLC2IOC"   // DB104
{ S7_Optimized_Access := 'FALSE' }
AUTHOR : KG
VERSION : 0.1
// Data sent to the IOC only to be used for communication between the PLC program and the IOC
   VAR
      HeartBeat : Word;
      Reserve : Array[0..37] of Byte;
   END_VAR
BEGIN
END_DATA_BLOCK

DATA_BLOCK "IOC2PLC"   // DB105
{ S7_Optimized_Access := 'FALSE' }
AUTHOR : KG
VERSION : 0.1
// Data to be sent from IOC to PLC. Used to send the information fromthe IOC tothe PLC (not for operator's commands)
   VAR
      HeartBeat : Word;
      TT900 : Real;
      TT930 : Real;
      TT940 : Real;
      TT950 : Real;
      TT960 : Real;
      TT630 : Real;
      TT640 : Real;
      TT700 : Real;
      TT650 : Real;
      TT660 : Real;
      TT610 : Real;
      TT620 : Real;
      TT600 : Real;
      TT670 : Real;
      TT680 : Real;
      TT690 : Real;
      TT970 : Real;
      TT980 : Real;
      TTf_VB_final1 : Real;
      TT06 : Real;
      TT07 : Real;
      "CTS:TT10" : Real;
      "CTS:TT11" : Real;
      "CTS:TT20" : Real;
      "CTS:TT21" : Real;
      TT04 : Real;
      TT05 : Real;
      "VBox:TT03" : Real;
      "CM:TT08" : Real;
      TT609 : Real;
      Reserved1 : Array[0..7] of Byte;
      TT900_VALID : Bool;
      TT930_VALID : Bool;
      TT940_VALID : Bool;
      TT950_VALID : Bool;
      TT960_VALID : Bool;
      TT630_VALID : Bool;
      TT640_VALID : Bool;
      TT700_VALID : Bool;
      TT650_VALID : Bool;
      TT660_VALID : Bool;
      TT610_VALID : Bool;
      TT620_VALID : Bool;
      TT600_VALID : Bool;
      TT670_VALID : Bool;
      TT680_VALID : Bool;
      TT690_VALID : Bool;
      TT970_VALID : Bool;
      TT980_VALID : Bool;
      TTf_VB_final1_VALID : Bool;
      TT06_VALID : Bool;
      TT07_VALID : Bool;
      "CTS:TT10_VALID" : Bool;
      "CTS:TT11_VALID" : Bool;
      "CTS:TT20_VALID" : Bool;
      "CTS:TT21_VALID" : Bool;
      TT04_VALID : Bool;
      TT05_VALID : Bool;
      "VBox:TT03_VALID" : Bool;
      "CM:TT08_VALID" : Bool;
      TT609_VALID : Bool;
      VALID_reserv6 : Bool;
      VALID_reserv7 : Bool;
      Reserved2 : Array[0..114] of Byte;
   END_VAR
BEGIN
END_DATA_BLOCK

DATA_BLOCK "S4_Parameters"   // DB204
TITLE = LN2 Screen cooling parameters
{ S7_Optimized_Access := 'FALSE' }
VERSION : 0.1
   VAR
      CV60_PID_GAIN : Real;
      CV60_PID_TI : Time;
      CV60_PID_TD : Time;
      CV60_PID_TM_LAG : Time;
      CV60_PID_LMN_HLM : Real;
      CV60_PID_LMN_LLM : Real;
      CV60_PID_SP_INT : Real;
   END_VAR
BEGIN
END_DATA_BLOCK

DATA_BLOCK "S6_parameters"   // DB206
{ S7_Optimized_Access := 'FALSE' }
VERSION : 0.1
   VAR
      CV02_PID_GAIN : Real;
      CV02_PID_TI : Time;
      CV02_PID_TD : Time;
      CV02_PID_TM_LAG : Time;
      CV03_PID_GAIN : Real;
      CV03_PID_TI : Time;
      CV03_PID_TD : Time;
      CV03_PID_TM_LAG : Time;
      TrigPID_CV02 : Real;
      PID_LT01_CV02_SP : Real;
      TrigPID_CV03 : Real;
      PID_LT03_CV03_SP : Real;
      PID_PT01_CV550_SP : Real;
      CV550 : Real;
      S5_P_FT552_MIN_GB : Real;
      S5_P_FT552_MAX_GB : Real;
      S5_P_FT552_MIN_C : Real;
      S5_P_FT552_MAX_C : Real;
   END_VAR
BEGIN
END_DATA_BLOCK

DATA_BLOCK "S7_Parameters"   // DB207
{ S7_Optimized_Access := 'FALSE' }
VERSION : 0.1
   VAR
      S7_LowT : Real;
      S7_HighT : Real;
   END_VAR
BEGIN
END_DATA_BLOCK

DATA_BLOCK "S8_parameters"   // DB208
{ S7_Optimized_Access := 'FALSE' }
AUTHOR : KG
VERSION : 0.1
   VAR
      CV01_Init : Real;
      CV01_open_rate : Real;
      "CM:TT08_cool" : Real;
      "VBox:TT03_cool" : Real;
      CV01_PID_GAIN : Real;
      CV01_PID_TI : Time;
      CV01_PID_TD : Time;
      CV01_PID_TM_LAG : Time;
      TrigPID_CV01 : Real;
      PID_LT01_CV01_SP : Real;
      S8_P_CV01 : Real;
      S8_P_CV01_Step7 : Real;
   END_VAR
BEGIN
END_DATA_BLOCK

DATA_BLOCK "#DATA_VALVES"   // DB306
TITLE = Instances of Valves
{ S7_Optimized_Access := 'FALSE' }
VERSION : 0.1
   VAR
      GV72 : "UDT_VALVES";
      RV90 : "UDT_VALVES";
      GV70 : "UDT_VALVES";
      Free_Valves : Array[0..3] of "UDT_VALVES";
   END_VAR
BEGIN
END_DATA_BLOCK

DATA_BLOCK "#DATA_HEATERS"   // DB313
{ S7_Optimized_Access := 'FALSE' }
VERSION : 0.1
// Heaters structures
   VAR
      EH90 : "UDT_HEATER";
      "EH93-96" : "UDT_HEATER";
      "EH63-70" : "UDT_HEATER";
      "EH61-62" : "UDT_HEATER";
      "EH60_67-69" : "UDT_HEATER";
      "EH97-98" : "UDT_HEATER";
      spareVB : Array[0..3] of "UDT_HEATER";
      EH01 : "UDT_HEATER";
      EH02 : "UDT_HEATER";
      EH10 : "UDT_HEATER";
      EH20 : "UDT_HEATER";
      "spare-CM-5" : "UDT_HEATER";
      "spare-CM-6" : "UDT_HEATER";
      "spare-CM-7" : "UDT_HEATER";
      "spare-CM-8" : "UDT_HEATER";
      "spare-CM-9" : "UDT_HEATER";
      "spare-CM-10" : "UDT_HEATER";
      "spare-CM-11" : "UDT_HEATER";
      "spare-CM-12" : "UDT_HEATER";
      EH12 : "UDT_HEATER";
      EH22 : "UDT_HEATER";
   END_VAR
BEGIN
END_DATA_BLOCK

// folder: SystemBlocksFolder/ReportSystemErrorFolder

DATA_BLOCK "RSE_DIAGNOSTIC_STATUS_DB"   // DB127
TITLE = Bloc de diagnostic Signalisation d'erreurs système
{ S7_Optimized_Access := 'FALSE' }
AUTHOR : SIMATIC
FAMILY : RSEDIAG
NAME : RSE7
VERSION : 1.0
// Ce DB fait partie de Signalisation d'erreurs système et sera actualisé par le FB de cette application.
//  Il constitue une interface pour la prise en charge du diagnostic système via la CPU serveur Web
   VAR
      Directory : Struct
      END_STRUCT;
      GlobalState : Struct
      END_STRUCT;
      Query : Struct
      END_STRUCT;
      Component : Struct
      END_STRUCT;
      Error : Struct
      END_STRUCT;
      State : Struct
      END_STRUCT;
      Alarm : Struct
      END_STRUCT;
      SubComponent : Struct
      END_STRUCT;
   END_VAR
BEGIN
END_DATA_BLOCK

// folder: (top level)

FUNCTION_BLOCK "graf"   // FB55, GRAPH
{ S7_Optimized_Access := 'FALSE' }
VERSION : 0.1
BEGIN